// TIA Portal project "uppgift2IndustriellIT" (V18) (continued)
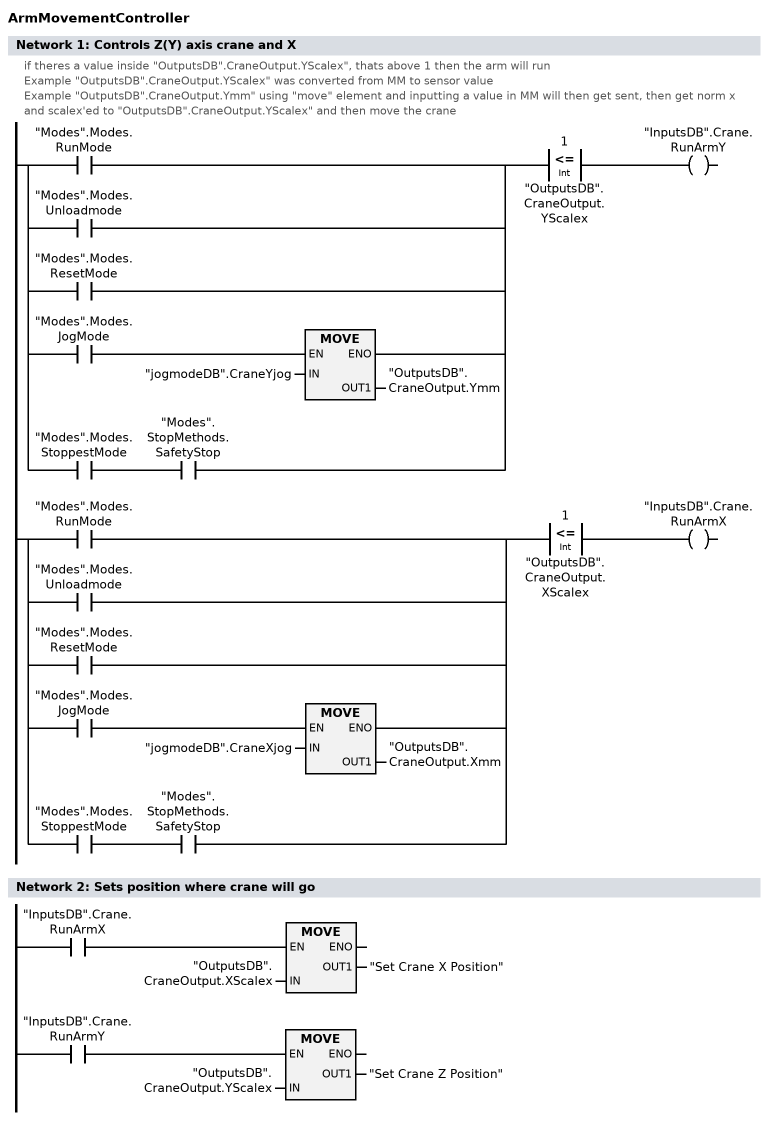
   RUNG wire#powerrail
      Contact( "Modes".Modes.RunMode )
      wire#w1
      { S7_Templates := "SrcType := Int" } LE_Contact(in1 := 1, in2 := "OutputsDB".CraneOutput.YScalex)
      Coil( "InputsDB".Crane.RunArmY )
   END_RUNG
   RUNG wire#powerrail
      Contact( "Modes".Modes.Unloadmode )
   END_RUNG wire#w1
   RUNG wire#powerrail
      Contact( "Modes".Modes.ResetMode )
   END_RUNG wire#w1
   RUNG wire#powerrail
      Contact( "Modes".Modes.JogMode )
      Move(in := "jogmodeDB".CraneYjog, out1 => "OutputsDB".CraneOutput.Ymm)
   END_RUNG wire#w1
   RUNG wire#powerrail
      Contact( "Modes".Modes.StoppestMode )
      Contact( "Modes".StopMethods.SafetyStop )
   END_RUNG wire#w1
   RUNG wire#powerrail
      Contact( "Modes".Modes.RunMode )
      wire#w2
      { S7_Templates := "SrcType := Int" } LE_Contact(in1 := 1, in2 := "OutputsDB".CraneOutput.XScalex)
      Coil( "InputsDB".Crane.RunArmX )
   END_RUNG
   RUNG wire#powerrail
      Contact( "Modes".Modes.Unloadmode )
   END_RUNG wire#w2
   RUNG wire#powerrail
      Contact( "Modes".Modes.ResetMode )
   END_RUNG wire#w2
   RUNG wire#powerrail
      Contact( "Modes".Modes.JogMode )
      Move(in := "jogmodeDB".CraneXjog, out1 => "OutputsDB".CraneOutput.Xmm)
   END_RUNG wire#w2
   RUNG wire#powerrail
      Contact( "Modes".Modes.StoppestMode )
      Contact( "Modes".StopMethods.SafetyStop )
   END_RUNG wire#w2
   // the same network as SCL:
   IF "Modes".Modes.JogMode THEN "OutputsDB".CraneOutput.Ymm := "jogmodeDB".CraneYjog; END_IF;
   "InputsDB".Crane.RunArmY := ("Modes".Modes.RunMode OR "Modes".Modes.Unloadmode OR "Modes".Modes.ResetMode OR "Modes".Modes.JogMode OR ("Modes".Modes.StoppestMode AND "Modes".StopMethods.SafetyStop)) AND (1 <= "OutputsDB".CraneOutput.YScalex);
   IF "Modes".Modes.JogMode THEN "OutputsDB".CraneOutput.Xmm := "jogmodeDB".CraneXjog; END_IF;
   "InputsDB".Crane.RunArmX := ("Modes".Modes.RunMode OR "Modes".Modes.Unloadmode OR "Modes".Modes.ResetMode OR "Modes".Modes.JogMode OR ("Modes".Modes.StoppestMode AND "Modes".StopMethods.SafetyStop)) AND (1 <= "OutputsDB".CraneOutput.XScalex);
END_REGION

REGION Network 2: Sets position where crane will go
   RUNG wire#powerrail
      Contact( "InputsDB".Crane.RunArmX )
      Move(in := "OutputsDB".CraneOutput.XScalex, out1 => "Set Crane X Position")
   END_RUNG
   RUNG wire#powerrail
      Contact( "InputsDB".Crane.RunArmY )
      Move(in := "OutputsDB".CraneOutput.YScalex, out1 => "Set Crane Z Position")
   END_RUNG
   // the same network as SCL:
   IF "InputsDB".Crane.RunArmX THEN "Set Crane X Position" := "OutputsDB".CraneOutput.XScalex; END_IF;
   IF "InputsDB".Crane.RunArmY THEN "Set Crane Z Position" := "OutputsDB".CraneOutput.YScalex; END_IF;
END_REGION
END_FUNCTION

FUNCTION "ArmCalibration" : Void   // FC12, SCL
{ S7_Optimized_Access := 'TRUE' }
VERSION : 0.1
BEGIN
   IF "HmiDb".HmiSaveArmCalX = TRUE AND "Modes".Modes.StoppestMode = TRUE THEN
       "PositionArray".XposCraneMM["HmiDb".XListColumn] := "HmiDb".CalInputVal;

   END_IF;

   IF "HmiDb".HmiSaveArmCalY = TRUE AND "Modes".Modes.StoppestMode = TRUE THEN
       "PositionArray".YposCraneMM["HmiDb".YListColumn] := "HmiDb".CalInputVal;

   END_IF;

   IF "InputsDB".PressAdjustX = TRUE THEN
       IF "InputsDB".AdjustX <= 0 THEN
           "jogmodeDB".CraneXjog := "jogmodeDB".CraneXjog + "InputsDB".AdjustX;
       ELSE
           "jogmodeDB".CraneXjog := "jogmodeDB".CraneXjog + "InputsDB".AdjustX;
       END_IF;
       "InputsDB".PressAdjustX := FALSE;
   END_IF;
   IF "InputsDB".PressAdjustY = TRUE THEN
       IF "InputsDB".AdjustY <= 0 THEN
           "jogmodeDB".CraneYjog := "jogmodeDB".CraneYjog + "InputsDB".AdjustY;
       ELSE
           "jogmodeDB".CraneYjog := "jogmodeDB".CraneYjog + "InputsDB".AdjustY;

       END_IF;
       "InputsDB".PressAdjustY := FALSE;
   END_IF;


   "HmiDb".CurrentPositionX := "PositionArray".XposCraneMM["HmiDb".XListColumn];
   "HmiDb".CurrentPositionY := "PositionArray".YposCraneMM["HmiDb".YListColumn];
END_FUNCTION

// folder: Functions/HmiRelatedFunc

FUNCTION "ConveyorCalibrater" : Void   // FC9, LAD
{ S7_Optimized_Access := 'TRUE' }
VERSION : 0.1
BEGIN

REGION Network 1: Depending on the chosen conveyor in calibration menu the HMI will show the saved values
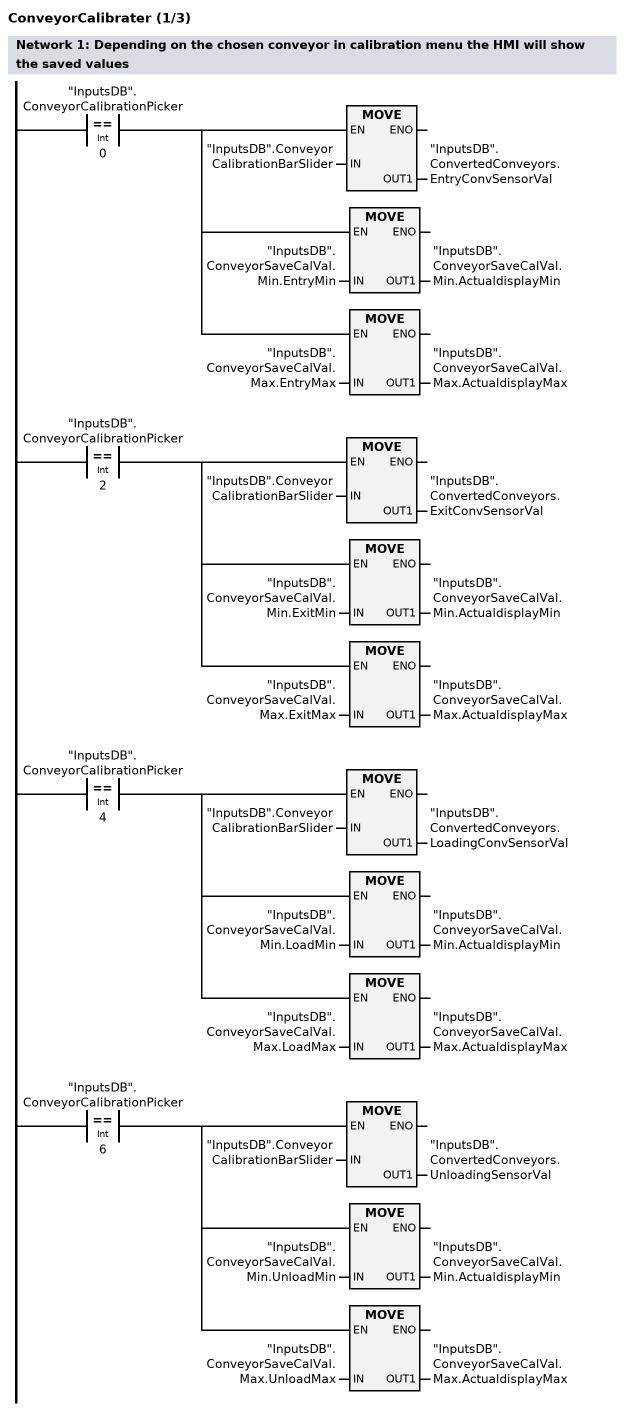
   RUNG wire#powerrail
      { S7_Templates := "SrcType := Int" } EQ_Contact(in1 := "InputsDB".ConveyorCalibrationPicker, in2 := 0)
      wire#w1
      Move(in := "InputsDB".ConveyorCalibrationBarSlider, out1 => "InputsDB".ConvertedConveyors.EntryConvSensorVal)
   END_RUNG
   RUNG wire#w1
      Move(in := "InputsDB".ConveyorSaveCalVal.Min.EntryMin, out1 => "InputsDB".ConveyorSaveCalVal.Min.ActualdisplayMin)
   END_RUNG
   RUNG wire#w1
      Move(in := "InputsDB".ConveyorSaveCalVal.Max.EntryMax, out1 => "InputsDB".ConveyorSaveCalVal.Max.ActualdisplayMax)
   END_RUNG
   RUNG wire#powerrail
      { S7_Templates := "SrcType := Int" } EQ_Contact(in1 := "InputsDB".ConveyorCalibrationPicker, in2 := 2)
      wire#w2
      Move(in := "InputsDB".ConveyorCalibrationBarSlider, out1 => "InputsDB".ConvertedConveyors.ExitConvSensorVal)
   END_RUNG
   RUNG wire#w2
      Move(in := "InputsDB".ConveyorSaveCalVal.Min.ExitMin, out1 => "InputsDB".ConveyorSaveCalVal.Min.ActualdisplayMin)
   END_RUNG
   RUNG wire#w2
      Move(in := "InputsDB".ConveyorSaveCalVal.Max.ExitMax, out1 => "InputsDB".ConveyorSaveCalVal.Max.ActualdisplayMax)
   END_RUNG
   RUNG wire#powerrail
      { S7_Templates := "SrcType := Int" } EQ_Contact(in1 := "InputsDB".ConveyorCalibrationPicker, in2 := 4)
      wire#w3
      Move(in := "InputsDB".ConveyorCalibrationBarSlider, out1 => "InputsDB".ConvertedConveyors.LoadingConvSensorVal)
   END_RUNG
   RUNG wire#w3
      Move(in := "InputsDB".ConveyorSaveCalVal.Min.LoadMin, out1 => "InputsDB".ConveyorSaveCalVal.Min.ActualdisplayMin)
   END_RUNG
   RUNG wire#w3
      Move(in := "InputsDB".ConveyorSaveCalVal.Max.LoadMax, out1 => "InputsDB".ConveyorSaveCalVal.Max.ActualdisplayMax)
   END_RUNG
   RUNG wire#powerrail
      { S7_Templates := "SrcType := Int" } EQ_Contact(in1 := "InputsDB".ConveyorCalibrationPicker, in2 := 6)
      wire#w4
      Move(in := "InputsDB".ConveyorCalibrationBarSlider, out1 => "InputsDB".ConvertedConveyors.UnloadingSensorVal)
   END_RUNG
   RUNG wire#w4
      Move(in := "InputsDB".ConveyorSaveCalVal.Min.UnloadMin, out1 => "InputsDB".ConveyorSaveCalVal.Min.ActualdisplayMin)
   END_RUNG
   RUNG wire#w4
      Move(in := "InputsDB".ConveyorSaveCalVal.Max.UnloadMax, out1 => "InputsDB".ConveyorSaveCalVal.Max.ActualdisplayMax)
   END_RUNG
   // the same network as SCL:
   IF "InputsDB".ConveyorCalibrationPicker = 0 THEN
       "InputsDB".ConvertedConveyors.EntryConvSensorVal := "InputsDB".ConveyorCalibrationBarSlider;
       "InputsDB".ConveyorSaveCalVal.Min.ActualdisplayMin := "InputsDB".ConveyorSaveCalVal.Min.EntryMin;
       "InputsDB".ConveyorSaveCalVal.Max.ActualdisplayMax := "InputsDB".ConveyorSaveCalVal.Max.EntryMax;
   END_IF;
   IF "InputsDB".ConveyorCalibrationPicker = 2 THEN
       "InputsDB".ConvertedConveyors.ExitConvSensorVal := "InputsDB".ConveyorCalibrationBarSlider;
       "InputsDB".ConveyorSaveCalVal.Min.ActualdisplayMin := "InputsDB".ConveyorSaveCalVal.Min.ExitMin;
       "InputsDB".ConveyorSaveCalVal.Max.ActualdisplayMax := "InputsDB".ConveyorSaveCalVal.Max.ExitMax;
   END_IF;
   IF "InputsDB".ConveyorCalibrationPicker = 4 THEN
       "InputsDB".ConvertedConveyors.LoadingConvSensorVal := "InputsDB".ConveyorCalibrationBarSlider;
       "InputsDB".ConveyorSaveCalVal.Min.ActualdisplayMin := "InputsDB".ConveyorSaveCalVal.Min.LoadMin;
       "InputsDB".ConveyorSaveCalVal.Max.ActualdisplayMax := "InputsDB".ConveyorSaveCalVal.Max.LoadMax;
   END_IF;
   IF "InputsDB".ConveyorCalibrationPicker = 6 THEN
       "InputsDB".ConvertedConveyors.UnloadingSensorVal := "InputsDB".ConveyorCalibrationBarSlider;
       "InputsDB".ConveyorSaveCalVal.Min.ActualdisplayMin := "InputsDB".ConveyorSaveCalVal.Min.UnloadMin;
       "InputsDB".ConveyorSaveCalVal.Max.ActualdisplayMax := "InputsDB".ConveyorSaveCalVal.Max.UnloadMax;
   END_IF;
END_REGION

REGION Network 2: saves the values from hmi
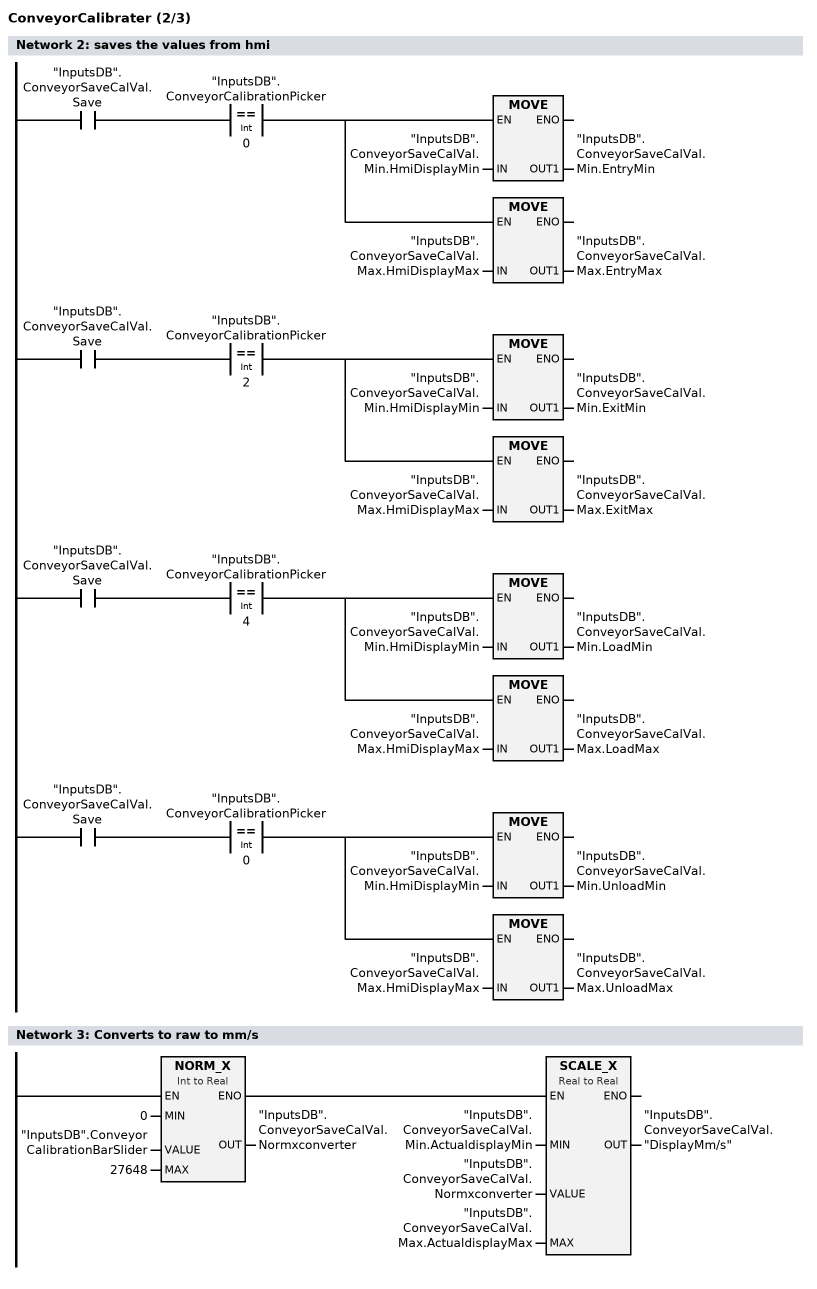
   RUNG wire#powerrail
      Contact( "InputsDB".ConveyorSaveCalVal.Save )
      { S7_Templates := "SrcType := Int" } EQ_Contact(in1 := "InputsDB".ConveyorCalibrationPicker, in2 := 0)
      wire#w1
      Move(in := "InputsDB".ConveyorSaveCalVal.Min.HmiDisplayMin, out1 => "InputsDB".ConveyorSaveCalVal.Min.EntryMin)
   END_RUNG
   RUNG wire#w1
      Move(in := "InputsDB".ConveyorSaveCalVal.Max.HmiDisplayMax, out1 => "InputsDB".ConveyorSaveCalVal.Max.EntryMax)
   END_RUNG
   RUNG wire#powerrail
      Contact( "InputsDB".ConveyorSaveCalVal.Save )
      { S7_Templates := "SrcType := Int" } EQ_Contact(in1 := "InputsDB".ConveyorCalibrationPicker, in2 := 2)
      wire#w2
      Move(in := "InputsDB".ConveyorSaveCalVal.Min.HmiDisplayMin, out1 => "InputsDB".ConveyorSaveCalVal.Min.ExitMin)
   END_RUNG
   RUNG wire#w2
      Move(in := "InputsDB".ConveyorSaveCalVal.Max.HmiDisplayMax, out1 => "InputsDB".ConveyorSaveCalVal.Max.ExitMax)
   END_RUNG
   RUNG wire#powerrail
      Contact( "InputsDB".ConveyorSaveCalVal.Save )
      { S7_Templates := "SrcType := Int" } EQ_Contact(in1 := "InputsDB".ConveyorCalibrationPicker, in2 := 4)
      wire#w3
      Move(in := "InputsDB".ConveyorSaveCalVal.Min.HmiDisplayMin, out1 => "InputsDB".ConveyorSaveCalVal.Min.LoadMin)
   END_RUNG
   RUNG wire#w3
      Move(in := "InputsDB".ConveyorSaveCalVal.Max.HmiDisplayMax, out1 => "InputsDB".ConveyorSaveCalVal.Max.LoadMax)
   END_RUNG
   RUNG wire#powerrail
      Contact( "InputsDB".ConveyorSaveCalVal.Save )
      { S7_Templates := "SrcType := Int" } EQ_Contact(in1 := "InputsDB".ConveyorCalibrationPicker, in2 := 0)
      wire#w4
      Move(in := "InputsDB".ConveyorSaveCalVal.Min.HmiDisplayMin, out1 => "InputsDB".ConveyorSaveCalVal.Min.UnloadMin)
   END_RUNG
   RUNG wire#w4
      Move(in := "InputsDB".ConveyorSaveCalVal.Max.HmiDisplayMax, out1 => "InputsDB".ConveyorSaveCalVal.Max.UnloadMax)
   END_RUNG
   // the same network as SCL:
   IF "InputsDB".ConveyorSaveCalVal.Save AND ("InputsDB".ConveyorCalibrationPicker = 0) THEN
       "InputsDB".ConveyorSaveCalVal.Min.EntryMin := "InputsDB".ConveyorSaveCalVal.Min.HmiDisplayMin;
       "InputsDB".ConveyorSaveCalVal.Max.EntryMax := "InputsDB".ConveyorSaveCalVal.Max.HmiDisplayMax;
   END_IF;
   IF "InputsDB".ConveyorSaveCalVal.Save AND ("InputsDB".ConveyorCalibrationPicker = 2) THEN
       "InputsDB".ConveyorSaveCalVal.Min.ExitMin := "InputsDB".ConveyorSaveCalVal.Min.HmiDisplayMin;
       "InputsDB".ConveyorSaveCalVal.Max.ExitMax := "InputsDB".ConveyorSaveCalVal.Max.HmiDisplayMax;
   END_IF;
   IF "InputsDB".ConveyorSaveCalVal.Save AND ("InputsDB".ConveyorCalibrationPicker = 4) THEN
       "InputsDB".ConveyorSaveCalVal.Min.LoadMin := "InputsDB".ConveyorSaveCalVal.Min.HmiDisplayMin;
       "InputsDB".ConveyorSaveCalVal.Max.LoadMax := "InputsDB".ConveyorSaveCalVal.Max.HmiDisplayMax;
   END_IF;
   IF "InputsDB".ConveyorSaveCalVal.Save AND ("InputsDB".ConveyorCalibrationPicker = 0) THEN
       "InputsDB".ConveyorSaveCalVal.Min.UnloadMin := "InputsDB".ConveyorSaveCalVal.Min.HmiDisplayMin;
       "InputsDB".ConveyorSaveCalVal.Max.UnloadMax := "InputsDB".ConveyorSaveCalVal.Max.HmiDisplayMax;
   END_IF;
END_REGION

REGION Network 3: Converts to raw to mm/s
   RUNG wire#powerrail
      { S7_Templates := "[SrcType := Int, DestType := Real]" } Normalize(min := 0, value := "InputsDB".ConveyorCalibrationBarSlider, max := 27648, out => "InputsDB".ConveyorSaveCalVal.Normxconverter)
      { S7_Templates := "[SrcType := Real, DestType := Real]" } Scale(min := "InputsDB".ConveyorSaveCalVal.Min.ActualdisplayMin, value := "InputsDB".ConveyorSaveCalVal.Normxconverter, max := "InputsDB".ConveyorSaveCalVal.Max.ActualdisplayMax, out => "InputsDB".ConveyorSaveCalVal."DisplayMm/s")
   END_RUNG
   // the same network as SCL:
   "InputsDB".ConveyorSaveCalVal.Normxconverter := NORM_X(MIN := 0, VALUE := "InputsDB".ConveyorCalibrationBarSlider, MAX := 27648);
   "InputsDB".ConveyorSaveCalVal."DisplayMm/s" := SCALE_X(MIN := "InputsDB".ConveyorSaveCalVal.Min.ActualdisplayMin, VALUE := "InputsDB".ConveyorSaveCalVal.Normxconverter, MAX := "InputsDB".ConveyorSaveCalVal.Max.ActualdisplayMax);
END_REGION

REGION Network 4: Prevents conveyor speed slider from being changed unless machine is stopped
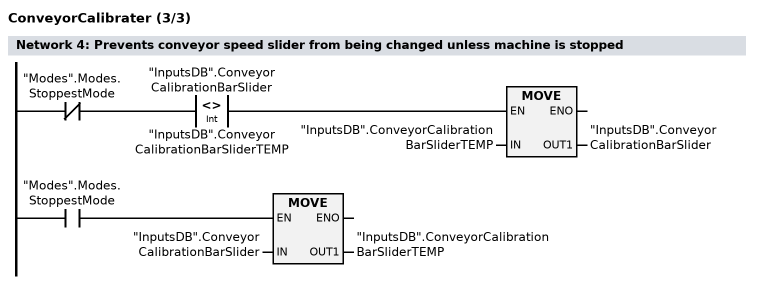
   RUNG wire#powerrail
      I_Contact( "Modes".Modes.StoppestMode )
      { S7_Templates := "SrcType := Int" } NE_Contact(in1 := "InputsDB".ConveyorCalibrationBarSlider, in2 := "InputsDB".ConveyorCalibrationBarSliderTEMP)
      Move(in := "InputsDB".ConveyorCalibrationBarSliderTEMP, out1 => "InputsDB".ConveyorCalibrationBarSlider)
   END_RUNG
   RUNG wire#powerrail
      Contact( "Modes".Modes.StoppestMode )
      Move(in := "InputsDB".ConveyorCalibrationBarSlider, out1 => "InputsDB".ConveyorCalibrationBarSliderTEMP)
   END_RUNG
   // the same network as SCL:
   IF NOT "Modes".Modes.StoppestMode AND ("InputsDB".ConveyorCalibrationBarSlider <> "InputsDB".ConveyorCalibrationBarSliderTEMP) THEN
       "InputsDB".ConveyorCalibrationBarSlider := "InputsDB".ConveyorCalibrationBarSliderTEMP;
   END_IF;
   IF "Modes".Modes.StoppestMode THEN
       "InputsDB".ConveyorCalibrationBarSliderTEMP := "InputsDB".ConveyorCalibrationBarSlider;
   END_IF;
END_REGION
END_FUNCTION

FUNCTION "Orders" : Void   // FC10, LAD
{ S7_Optimized_Access := 'TRUE' }
VERSION : 0.1
   VAR_TEMP   // added for the SCL form of the ladder/FBD networks
      _w1 : Bool;
   END_VAR
BEGIN

REGION Network 1: Enables order mode
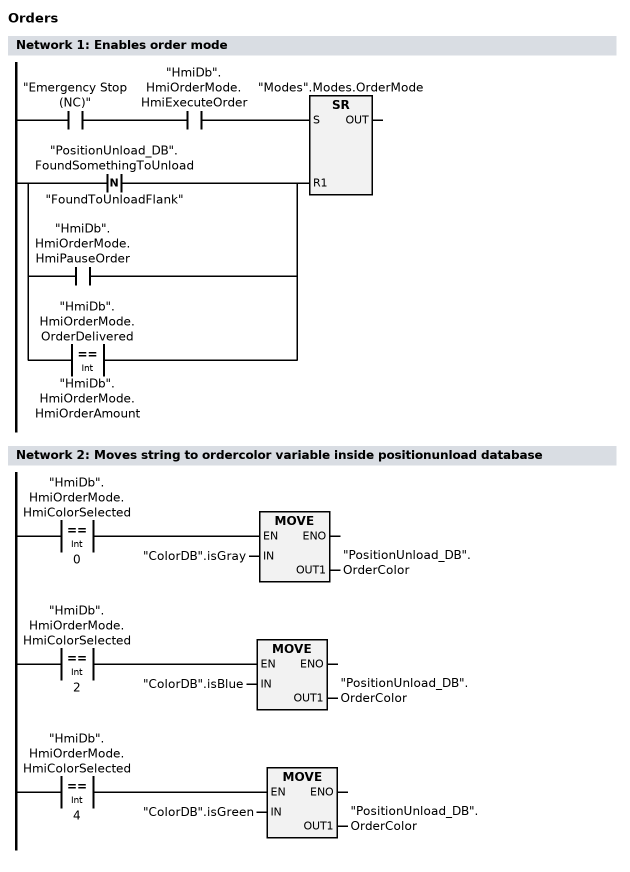
   RUNG wire#powerrail
      Contact( "Emergency Stop (NC)" )
      Contact( "HmiDb".HmiOrderMode.HmiExecuteOrder )
      S_SR(operand := "Modes".Modes.OrderMode, r1 := wire#w1)
   END_RUNG
   RUNG wire#powerrail
      N_Contact(operand := "PositionUnload_DB".FoundSomethingToUnload, bit := "FoundToUnloadFlank")
   END_RUNG wire#w1
   RUNG wire#powerrail
      Contact( "HmiDb".HmiOrderMode.HmiPauseOrder )
   END_RUNG wire#w1
   RUNG wire#powerrail
      { S7_Templates := "SrcType := Int" } EQ_Contact(in1 := "HmiDb".HmiOrderMode.OrderDelivered, in2 := "HmiDb".HmiOrderMode.HmiOrderAmount)
   END_RUNG wire#w1
   // the same network as SCL:
   #_w1 := NOT "PositionUnload_DB".FoundSomethingToUnload AND "FoundToUnloadFlank";   // falling edge of "PositionUnload_DB".FoundSomethingToUnload
   "FoundToUnloadFlank" := "PositionUnload_DB".FoundSomethingToUnload;
   IF "Emergency Stop (NC)" AND "HmiDb".HmiOrderMode.HmiExecuteOrder THEN
       "Modes".Modes.OrderMode := TRUE;   // SR flip-flop
   END_IF;
   IF #_w1 OR "HmiDb".HmiOrderMode.HmiPauseOrder OR ("HmiDb".HmiOrderMode.OrderDelivered = "HmiDb".HmiOrderMode.HmiOrderAmount) THEN
       "Modes".Modes.OrderMode := FALSE;
   END_IF;
END_REGION

REGION Network 2: Moves string to ordercolor variable inside positionunload database
   RUNG wire#powerrail
      { S7_Templates := "SrcType := Int" } EQ_Contact(in1 := "HmiDb".HmiOrderMode.HmiColorSelected, in2 := 0)
      Move(in := "ColorDB".isGray, out1 => "PositionUnload_DB".OrderColor)
   END_RUNG
   RUNG wire#powerrail
      { S7_Templates := "SrcType := Int" } EQ_Contact(in1 := "HmiDb".HmiOrderMode.HmiColorSelected, in2 := 2)
      Move(in := "ColorDB".isBlue, out1 => "PositionUnload_DB".OrderColor)
   END_RUNG
   RUNG wire#powerrail
      { S7_Templates := "SrcType := Int" } EQ_Contact(in1 := "HmiDb".HmiOrderMode.HmiColorSelected, in2 := 4)
      Move(in := "ColorDB".isGreen, out1 => "PositionUnload_DB".OrderColor)
   END_RUNG
   // the same network as SCL:
   IF "HmiDb".HmiOrderMode.HmiColorSelected = 0 THEN
       "PositionUnload_DB".OrderColor := "ColorDB".isGray;
   END_IF;
   IF "HmiDb".HmiOrderMode.HmiColorSelected = 2 THEN
       "PositionUnload_DB".OrderColor := "ColorDB".isBlue;
   END_IF;
   IF "HmiDb".HmiOrderMode.HmiColorSelected = 4 THEN
       "PositionUnload_DB".OrderColor := "ColorDB".isGreen;
   END_IF;
END_REGION
END_FUNCTION

FUNCTION "HmiAnimations" : Void   // FC11, LAD
{ S7_Optimized_Access := 'TRUE' }
VERSION : 0.1
BEGIN

REGION Network 1: changevalue to move box animation in hmi
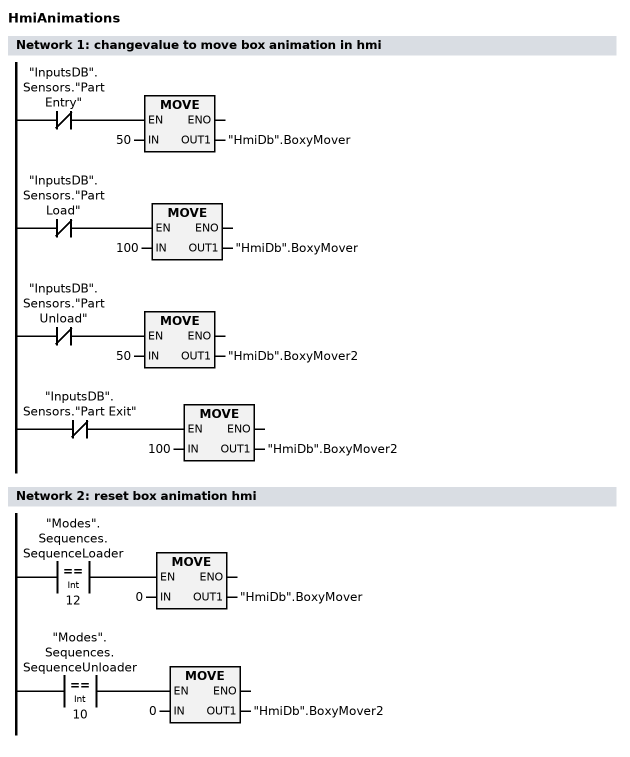
   RUNG wire#powerrail
      I_Contact( "InputsDB".Sensors."Part Entry" )
      Move(in := 50, out1 => "HmiDb".BoxyMover)
   END_RUNG
   RUNG wire#powerrail
      I_Contact( "InputsDB".Sensors."Part Load" )
      Move(in := 100, out1 => "HmiDb".BoxyMover)
   END_RUNG
   RUNG wire#powerrail
      I_Contact( "InputsDB".Sensors."Part Unload" )
      Move(in := 50, out1 => "HmiDb".BoxyMover2)
   END_RUNG
   RUNG wire#powerrail
      I_Contact( "InputsDB".Sensors."Part Exit" )
      Move(in := 100, out1 => "HmiDb".BoxyMover2)
   END_RUNG
   // the same network as SCL:
   IF NOT "InputsDB".Sensors."Part Entry" THEN "HmiDb".BoxyMover := 50; END_IF;
   IF NOT "InputsDB".Sensors."Part Load" THEN "HmiDb".BoxyMover := 100; END_IF;
   IF NOT "InputsDB".Sensors."Part Unload" THEN "HmiDb".BoxyMover2 := 50; END_IF;
   IF NOT "InputsDB".Sensors."Part Exit" THEN "HmiDb".BoxyMover2 := 100; END_IF;
END_REGION

REGION Network 2: reset box animation hmi
   RUNG wire#powerrail
      { S7_Templates := "SrcType := Int" } EQ_Contact(in1 := "Modes".Sequences.SequenceLoader, in2 := 12)
      Move(in := 0, out1 => "HmiDb".BoxyMover)
   END_RUNG
   RUNG wire#powerrail
      { S7_Templates := "SrcType := Int" } EQ_Contact(in1 := "Modes".Sequences.SequenceUnloader, in2 := 10)
      Move(in := 0, out1 => "HmiDb".BoxyMover2)
   END_RUNG
   // the same network as SCL:
   IF "Modes".Sequences.SequenceLoader = 12 THEN "HmiDb".BoxyMover := 0; END_IF;
   IF "Modes".Sequences.SequenceUnloader = 10 THEN "HmiDb".BoxyMover2 := 0; END_IF;
END_REGION
END_FUNCTION

// folder: Functions/SCL

FUNCTION_BLOCK "PositionsLoad"   // FB1, SCL
{ S7_Optimized_Access := 'TRUE' }
VERSION : 0.1
   VAR_INPUT
      debouncer : Int;
      index : Int;
      index2 : Int := 0;
      FoundEmpty : Bool;
      roww : Int := 0;
      VisionSensorVal : Int;
      yas : Int;
   END_VAR
BEGIN
   IF "Modes".Sequences.SequenceLoader = 13 AND "Modes".Modes.StoppestMode = FALSE THEN
       FOR #index := 0 TO 5 DO
           IF #debouncer = 0 THEN //Om inte existerar kommer for loopen att köras klart innan armen hinner göra något
               #FoundEmpty := FALSE;

               IF "AlreadyFilledSlotArray".Row1Y[#index] = 0 THEN
                   #debouncer := 1;

                   "OutputsDB".CraneOutput.Ymm := "PositionArray".YposCraneMM[#index];
                   "OutputsDB".CraneOutput.Xmm := "PositionArray".XposCraneMM[#index2];
                   #FoundEmpty := TRUE;
                   "AlreadyFilledSlotArray".Row1Y[#index] := #VisionSensorVal;
                   EXIT;
               END_IF;

               IF "AlreadyFilledSlotArray".Row2Y[#index] = 0 THEN
                   #debouncer := 1;
                   "AlreadyFilledSlotArray".Row2Y[#index] := #VisionSensorVal;
                   "OutputsDB".CraneOutput.Ymm := "PositionArray".YposCraneMM[#index];
                   "OutputsDB".CraneOutput.Xmm := "PositionArray".XposCraneMM[#index2 + 1];
                   #FoundEmpty := TRUE;
                   EXIT;
               END_IF;
               IF "AlreadyFilledSlotArray".Row3Y[#index] = 0 THEN
                   #debouncer := 1;
                   "AlreadyFilledSlotArray".Row3Y[#index] := #VisionSensorVal;
                   "OutputsDB".CraneOutput.Ymm := "PositionArray".YposCraneMM[#index];
                   "OutputsDB".CraneOutput.Xmm := "PositionArray".XposCraneMM[#index2 + 2];
                   #FoundEmpty := TRUE;
                   EXIT;
               END_IF;
               IF "AlreadyFilledSlotArray".Row4Y[#index] = 0 THEN
                   #debouncer := 1;
                   "AlreadyFilledSlotArray".Row4Y[#index] := #VisionSensorVal;
                   "OutputsDB".CraneOutput.Ymm := "PositionArray".YposCraneMM[#index];
                   "OutputsDB".CraneOutput.Xmm := "PositionArray".XposCraneMM[#index2 + 3];
                   #FoundEmpty := TRUE;
                   EXIT;

               END_IF;

               IF "AlreadyFilledSlotArray".Row5Y[#index] = 0 THEN
                   #debouncer := 1;
                   "AlreadyFilledSlotArray".Row5Y[#index] := #VisionSensorVal;
                   "OutputsDB".CraneOutput.Ymm := "PositionArray".YposCraneMM[#index];
                   "OutputsDB".CraneOutput.Xmm := "PositionArray".XposCraneMM[#index2 + 4];
                   #FoundEmpty := TRUE;
                   EXIT;
               END_IF;
               IF "AlreadyFilledSlotArray".Row6Y[#index] = 0 THEN
                   #debouncer := 1;
                   "AlreadyFilledSlotArray".Row6Y[#index] := #VisionSensorVal;
                   "OutputsDB".CraneOutput.Ymm := "PositionArray".YposCraneMM[#index];
                   "OutputsDB".CraneOutput.Xmm := "PositionArray".XposCraneMM[#index2 + 5];
                   #FoundEmpty := TRUE;
                   EXIT;
               END_IF;
               IF "AlreadyFilledSlotArray".Row7Y[#index] = 0 THEN
                   #debouncer := 1;
                   "AlreadyFilledSlotArray".Row7Y[#index] := #VisionSensorVal;
                   "OutputsDB".CraneOutput.Ymm := "PositionArray".YposCraneMM[#index];
                   "OutputsDB".CraneOutput.Xmm := "PositionArray".XposCraneMM[#index2 + 6];
                   #FoundEmpty := TRUE;
                   EXIT;

               END_IF;
               IF "AlreadyFilledSlotArray".Row8Y[#index] = 0 THEN
                   #debouncer := 1;
                   "AlreadyFilledSlotArray".Row8Y[#index] := #VisionSensorVal;
                   "OutputsDB".CraneOutput.Ymm := "PositionArray".YposCraneMM[#index];
                   "OutputsDB".CraneOutput.Xmm := "PositionArray".XposCraneMM[#index2 + 7];
                   #FoundEmpty := TRUE;
                   EXIT;
               END_IF;
               IF "AlreadyFilledSlotArray".Row9Y[#index] = 0 THEN
                   #debouncer := 1;
                   "AlreadyFilledSlotArray".Row9Y[#index] := #VisionSensorVal;
                   "OutputsDB".CraneOutput.Ymm := "PositionArray".YposCraneMM[#index];
                   "OutputsDB".CraneOutput.Xmm := "PositionArray".XposCraneMM[#index2 + 8];
                   #FoundEmpty := TRUE;
                   EXIT;
               END_IF;


           END_IF;

       END_FOR;
       IF #FoundEmpty = FALSE THEN
           "Modes".Modes.StoppestMode := TRUE;
       END_IF;


   END_IF;
END_FUNCTION_BLOCK

FUNCTION_BLOCK "PositionUnload"   // FB2, SCL
{ S7_Optimized_Access := 'TRUE' }
VERSION : 0.1
   VAR_INPUT
      index : Int;
      index2 : Int;
      debouncer : Int;
      FoundSomethingToUnload : Bool;
      OrderColor : Int;
      ColorUnloaded : Int;
   END_VAR
BEGIN

   FOR #index := 0 TO 5 DO
       IF #debouncer = 0 THEN
           #FoundSomethingToUnload := FALSE; //ifall false innebär ifall for loopen körs klart och den inte blir true innebär att lagret är tomt
           IF "AlreadyFilledSlotArray".Row1Y[#index] <> 0 THEN
               #FoundSomethingToUnload := TRUE; //hittade något att lasta ut
               IF "Modes".Modes.OrderMode = TRUE THEN //om order mode aktiv
                   IF "AlreadyFilledSlotArray".Row1Y[#index] = #OrderColor THEN //Om hittade färgen som användaren ville unloada
                       #debouncer := 1; //aktiverar debouncern
                       "AlreadyFilledSlotArray".Row1Y[#index] := 0; //Uppdaterar db
                       "OutputsDB".CraneOutput.Ymm := "PositionArray".YposCraneMM[#index];
                       "OutputsDB".CraneOutput.Xmm := "PositionArray".XposCraneMM[#index2];
                       EXIT;
                   END_IF;

               END_IF;
               IF "Modes".Modes.OrderMode = FALSE THEN
                   #debouncer := 1;
                   #ColorUnloaded := "AlreadyFilledSlotArray".Row1Y[#index];
                   "AlreadyFilledSlotArray".Row1Y[#index] := 0;
                   "OutputsDB".CraneOutput.Ymm := "PositionArray".YposCraneMM[#index];
                   "OutputsDB".CraneOutput.Xmm := "PositionArray".XposCraneMM[#index2];

                   EXIT;
               END_IF;
           END_IF;

           //yessssssssssssssssssssssss

           IF "AlreadyFilledSlotArray".Row2Y[#index] <> 0 THEN
               #FoundSomethingToUnload := TRUE;
               IF "Modes".Modes.OrderMode = TRUE THEN
                   IF "AlreadyFilledSlotArray".Row2Y[#index] = #OrderColor THEN

                       #debouncer := 1;

                       "AlreadyFilledSlotArray".Row2Y[#index] := 0;
                       "OutputsDB".CraneOutput.Ymm := "PositionArray".YposCraneMM[#index];
                       "OutputsDB".CraneOutput.Xmm := "PositionArray".XposCraneMM[#index2+1];
                       EXIT;
                   END_IF
                   ;
               END_IF;
               IF "Modes".Modes.OrderMode = FALSE THEN
                   #debouncer := 1;
                   #ColorUnloaded := "AlreadyFilledSlotArray".Row2Y[#index];
                   "AlreadyFilledSlotArray".Row2Y[#index] := 0;
                   "OutputsDB".CraneOutput.Ymm := "PositionArray".YposCraneMM[#index];
                   "OutputsDB".CraneOutput.Xmm := "PositionArray".XposCraneMM[#index2 + 1];

                   EXIT;
               END_IF;
               END_IF;

               //yessssssssssssssssssssssss
               //

               IF "AlreadyFilledSlotArray".Row3Y[#index] <> 0 THEN
                   #FoundSomethingToUnload := TRUE;
                   IF "Modes".Modes.OrderMode = TRUE THEN
                       IF "AlreadyFilledSlotArray".Row3Y[#index] = #OrderColor THEN

                           #debouncer := 1;

                           "AlreadyFilledSlotArray".Row3Y[#index] := 0;
                           "OutputsDB".CraneOutput.Ymm := "PositionArray".YposCraneMM[#index];
                           "OutputsDB".CraneOutput.Xmm := "PositionArray".XposCraneMM[#index2 + 2];
                           EXIT;
                       END_IF
                       ;
                   END_IF;
                   IF "Modes".Modes.OrderMode = FALSE THEN
                       #debouncer := 1;
                       #ColorUnloaded := "AlreadyFilledSlotArray".Row3Y[#index];
                       "AlreadyFilledSlotArray".Row3Y[#index] := 0;
                       "OutputsDB".CraneOutput.Ymm := "PositionArray".YposCraneMM[#index];
                       "OutputsDB".CraneOutput.Xmm := "PositionArray".XposCraneMM[#index2 + 2];

                       EXIT;
                   END_IF;
               END_IF;

               //yessssssssssssssssssssssss
               //


               IF "AlreadyFilledSlotArray".Row4Y[#index] <> 0 THEN
                   #FoundSomethingToUnload := TRUE;
                   IF "Modes".Modes.OrderMode = TRUE THEN
                       IF "AlreadyFilledSlotArray".Row4Y[#index] = #OrderColor THEN

                           #debouncer := 1;

                           "AlreadyFilledSlotArray".Row4Y[#index] := 0;
                           "OutputsDB".CraneOutput.Ymm := "PositionArray".YposCraneMM[#index];
                           "OutputsDB".CraneOutput.Xmm := "PositionArray".XposCraneMM[#index2 + 3];
                           EXIT;
                       END_IF
                       ;
                   END_IF;
                   IF "Modes".Modes.OrderMode = FALSE THEN
                       #ColorUnloaded := "AlreadyFilledSlotArray".Row4Y[#index];
                       #debouncer := 1;
                       "AlreadyFilledSlotArray".Row4Y[#index] := 0;
                       "OutputsDB".CraneOutput.Ymm := "PositionArray".YposCraneMM[#index];
                       "OutputsDB".CraneOutput.Xmm := "PositionArray".XposCraneMM[#index2 + 3];

                       EXIT;
                   END_IF;
               END_IF;

               //yessssssssssssssssssssssss
               //
               IF "AlreadyFilledSlotArray".Row5Y[#index] <> 0 THEN
                   #FoundSomethingToUnload := TRUE;
                   IF "Modes".Modes.OrderMode = TRUE THEN
                       IF "AlreadyFilledSlotArray".Row5Y[#index] = #OrderColor THEN

                           #debouncer := 1;

                           "AlreadyFilledSlotArray".Row5Y[#index] := 0;
                           "OutputsDB".CraneOutput.Ymm := "PositionArray".YposCraneMM[#index];
                           "OutputsDB".CraneOutput.Xmm := "PositionArray".XposCraneMM[#index2 + 4];
                           EXIT;
                       END_IF
                       ;
                   END_IF;
                   IF "Modes".Modes.OrderMode = FALSE THEN
                       #debouncer := 1;
                       #ColorUnloaded := "AlreadyFilledSlotArray".Row5Y[#index];
                       "AlreadyFilledSlotArray".Row5Y[#index] := 0;
                       "OutputsDB".CraneOutput.Ymm := "PositionArray".YposCraneMM[#index];
                       "OutputsDB".CraneOutput.Xmm := "PositionArray".XposCraneMM[#index2 + 4];

                       EXIT;
                   END_IF;
               END_IF;

               IF "AlreadyFilledSlotArray".Row6Y[#index] <> 0 THEN
                   #FoundSomethingToUnload := TRUE;
                   IF "Modes".Modes.OrderMode = TRUE THEN
                       IF "AlreadyFilledSlotArray".Row6Y[#index] = #OrderColor THEN

                           #debouncer := 1;

                           "AlreadyFilledSlotArray".Row6Y[#index] := 0;
                           "OutputsDB".CraneOutput.Ymm := "PositionArray".YposCraneMM[#index];
                           "OutputsDB".CraneOutput.Xmm := "PositionArray".XposCraneMM[#index2 + 5];
                           EXIT;
                       END_IF
                       ;
                   END_IF;
                   IF "Modes".Modes.OrderMode = FALSE THEN
                       #debouncer := 1;
                       #ColorUnloaded := "AlreadyFilledSlotArray".Row6Y[#index];
                       "AlreadyFilledSlotArray".Row6Y[#index] := 0;

                       "OutputsDB".CraneOutput.Ymm := "PositionArray".YposCraneMM[#index];
                       "OutputsDB".CraneOutput.Xmm := "PositionArray".XposCraneMM[#index2 + 5];

                       EXIT;
                   END_IF;
               END_IF;
               //yesssssssssssssss
               //

               IF "AlreadyFilledSlotArray".Row7Y[#index] <> 0 THEN
                   #FoundSomethingToUnload := TRUE;
                   IF "Modes".Modes.OrderMode = TRUE THEN
                       IF "AlreadyFilledSlotArray".Row7Y[#index] = #OrderColor THEN

                           #debouncer := 1;

                           "AlreadyFilledSlotArray".Row7Y[#index] := 0;
                           "OutputsDB".CraneOutput.Ymm := "PositionArray".YposCraneMM[#index];
                           "OutputsDB".CraneOutput.Xmm := "PositionArray".XposCraneMM[#index2 + 6];
                           EXIT;
                       END_IF
                       ;
                   END_IF;
                   IF "Modes".Modes.OrderMode = FALSE THEN
                       #debouncer := 1;
                       #ColorUnloaded := "AlreadyFilledSlotArray".Row7Y[#index];

                       "AlreadyFilledSlotArray".Row7Y[#index] := 0;
                       "OutputsDB".CraneOutput.Ymm := "PositionArray".YposCraneMM[#index];
                       "OutputsDB".CraneOutput.Xmm := "PositionArray".XposCraneMM[#index2 + 6];

                       EXIT;
                   END_IF;
               END_IF;
               //yesssssssssssssss
               //
               IF "AlreadyFilledSlotArray".Row8Y[#index] <> 0 THEN
                   #FoundSomethingToUnload := TRUE;
                   IF "Modes".Modes.OrderMode = TRUE THEN
                       IF "AlreadyFilledSlotArray".Row8Y[#index] = #OrderColor THEN

                           #debouncer := 1;

                           "AlreadyFilledSlotArray".Row8Y[#index] := 0;
                           "OutputsDB".CraneOutput.Ymm := "PositionArray".YposCraneMM[#index];
                           "OutputsDB".CraneOutput.Xmm := "PositionArray".XposCraneMM[#index2 + 7];
                           EXIT;
                       END_IF
                       ;
                   END_IF;
                   IF "Modes".Modes.OrderMode = FALSE THEN
                       #debouncer := 1;
                       #ColorUnloaded := "AlreadyFilledSlotArray".Row8Y[#index];
                       "AlreadyFilledSlotArray".Row8Y[#index] := 0;
                       "OutputsDB".CraneOutput.Ymm := "PositionArray".YposCraneMM[#index];
                       "OutputsDB".CraneOutput.Xmm := "PositionArray".XposCraneMM[#index2 + 7];

                       EXIT;
                   END_IF;
               END_IF;
               //yesssssssssssssss
               //
               IF "AlreadyFilledSlotArray".Row9Y[#index] <> 0 THEN
                   #FoundSomethingToUnload := TRUE;
                   IF "Modes".Modes.OrderMode = TRUE THEN
                       IF "AlreadyFilledSlotArray".Row9Y[#index] = #OrderColor THEN

                           #debouncer := 1;

                           "AlreadyFilledSlotArray".Row9Y[#index] := 0;
                           "OutputsDB".CraneOutput.Ymm := "PositionArray".YposCraneMM[#index];
                           "OutputsDB".CraneOutput.Xmm := "PositionArray".XposCraneMM[#index2 + 8];
                           EXIT;
                       END_IF
                       ;
                   END_IF;
                   IF "Modes".Modes.OrderMode = FALSE THEN
                       #debouncer := 1;
                       #ColorUnloaded := "AlreadyFilledSlotArray".Row9Y[#index];
                       "AlreadyFilledSlotArray".Row9Y[#index] := 0;
                       "OutputsDB".CraneOutput.Ymm := "PositionArray".YposCraneMM[#index];
                       "OutputsDB".CraneOutput.Xmm := "PositionArray".XposCraneMM[#index2 + 8];

                       EXIT;
                   END_IF;
               END_IF;
               //yesssssssssssssss
               //
       END_IF;


   END_FOR;


   IF #FoundSomethingToUnload = FALSE AND "Modes".Modes.OrderMode = FALSE THEN
       "Modes".Modes.StoppestMode := TRUE;
   END_IF;

   IF #FoundSomethingToUnload = FALSE AND "Modes".Modes.OrderMode = TRUE THEN
       "Modes".Modes.OrderMode := FALSE;
   END_IF;
END_FUNCTION_BLOCK

FUNCTION_BLOCK "resetFill"   // FB3, SCL
{ S7_Optimized_Access := 'TRUE' }
VERSION : 0.1
   VAR_INPUT
      i : Int;
   END_VAR
BEGIN
       FOR #i := 0 TO 5 DO
           "AlreadyFilledSlotArray".Row1Y[#i] := 0;
           "AlreadyFilledSlotArray".Row2Y[#i] := 0;
           "AlreadyFilledSlotArray".Row3Y[#i] := 0;
           "AlreadyFilledSlotArray".Row4Y[#i] := 0;
           "AlreadyFilledSlotArray".Row5Y[#i] := 0;
           "AlreadyFilledSlotArray".Row6Y[#i] := 0;
           "AlreadyFilledSlotArray".Row7Y[#i] := 0;
           "AlreadyFilledSlotArray".Row8Y[#i] := 0;
           "AlreadyFilledSlotArray".Row9Y[#i] := 0;
       END_FOR;
END_FUNCTION_BLOCK

// folder: Functions/input/output

FUNCTION "Inputs" : Void   // FC3, LAD
{ S7_Optimized_Access := 'TRUE' }
VERSION : 0.1
   VAR_TEMP   // added for the SCL form of the ladder/FBD networks
      _w1 : Bool;
      _w2 : Bool;
      _w3 : Bool;
   END_VAR
BEGIN

REGION Network 1: Set the modes (run mode, stop mode, reset mode)
   // Resetmode innehåller även visionsensor felhantering, resetmode sekvensen är i Outputs funktionen